screen "Dos" 800x480, template "Main"
   Group "Group_1" at 127,146 size 416x126; Text 'Мешалка 1'; PictureList "Motor"; TextList "Hand"; Picture "z2use_3"
   Group "Group_2" at 127,285 size 416x126; Text 'Мешалка 1'; PictureList "Motor"; TextList "Hand"; Picture "z2use_3"
   Rectangle "Rectangle_1" at 127,7 size 416x126
      Appearance <- "Motors_DB_M1_CMD_Sim"
   GraphicIOField "Graphic I/O field_2" at 134,43 size 43x85; PictureList "Motor"
      ProcessValue <- "Motors_DB_M1_Status"
   Button "Button_7" at 213,41 size 90x22; TextOff 'Авто'; TextList "Hand"
      on Click: InvertBit("Motors_DB_M1_CMD_Hand")
      Appearance <- "Motors_DB_M1_CMD_Hand"
      ProcessValue <- "Motors_DB_M1_CMD_Hand"
   Button "Button_8" at 258,63 size 45x22; TextOff 'Выкл'
      on Click: ResetBit("Motors_DB_M1_CMD_Start_M")
   Button "Button_9" at 213,86 size 90x20; TextOff 'Сервис'
      on Click: InvertBit("Motors_DB_M1_CMD_Service")
      Appearance <- "Motors_DB_M1_CMD_Service"
   Button "Button_13" at 213,63 size 45x22; TextOff 'Вкл'
      on Click: SetBit("Motors_DB_M1_CMD_Start_M")
      Appearance <- "Motors_DB_M1_CMD_Start_M"
   TextField "Text field_13" at 133,12 size 171x26; Text 'Дозатор 1'
   TextField "Text field_15" at 310,12 size 99x18; Text 'Ожидание ОС, с'
   GraphicView "Graphic view_1" at 180,42 size 25x25; Picture "z2use_3"
      Visibility <- "Motors_DB_M1_CMD_Hand"
   GraphicView "Graphic view_8" at 180,74 size 25x25; Picture "force"
      Visibility <- "Motors_DB_M1_CMD_Force"
   GraphicView "Graphic view_11" at 180,103 size 25x25; Picture "service"
      Visibility <- "Motors_DB_M1_CMD_Service"
   TextField "Text field_3" at 436,31 size 20x18; Text 'QF'
   TextField "Text field_10" at 436,56 size 21x18; Text 'KM'
   TextField "Text field_12" at 436,82 size 44x18; Text 'Service'
   TextField "Text field_14" at 436,108 size 41x18; Text 'Termo'
   TextField "Text field_4" at 416,10 size 120x22; Text 'Использовать:'
   Button "Button_21" at 478,32 size 60x20; TextOff 'Text'; Authorization "Operator"; PictureList "ON_OFF"
      on Click: InvertBit("Motors_DB_M1_Use_QF")
      ProcessValue <- "Motors_DB_M1_Use_QF"
   Button "Button_22" at 478,56 size 60x20; TextOff 'Text'; PictureList "ON_OFF"; Authorization "Operator"
      on Click: InvertBit("Motors_DB_M1_Use_KM")
      ProcessValue <- "Motors_DB_M1_Use_KM"
   Button "Button_24" at 478,80 size 60x20; TextOff 'Text'; PictureList "ON_OFF"; Authorization "Operator"
      on Click: InvertBit("Motors_DB_M1_Use_Serivce")
      ProcessValue <- "Motors_DB_M1_Use_Serivce"
   Button "Button_25" at 478,105 size 60x20; TextOff 'Text'; PictureList "ON_OFF"; Authorization "Operator"
      on Click: InvertBit("Motors_DB_M1_Use_Termo")
      ProcessValue <- "Motors_DB_M1_Use_Termo"
   Button "Button_26" at 416,31 size 20x20; TextOff 'Text'; Authorization "Operator"; PictureList "ok"
      ProcessValue <- "Motors_DB_M1_FB_QF"
   Button "Button_27" at 416,55 size 20x20; TextOff 'Text'; PictureList "ok"; Authorization "Operator"
      ProcessValue <- "Motors_DB_M1_FB_KM"
   Button "Button_29" at 416,80 size 20x20; TextOff 'Text'; PictureList "ok"; Authorization "Operator"
      ProcessValue <- "Motors_DB_M1_Use_Serivce"
   Button "Button_30" at 416,105 size 20x20; TextOff 'Text'; PictureList "ok"; Authorization "Operator"
      ProcessValue <- "Motors_DB_M1_FB_Termo"
   TextField "Text field_1" at 323,87 size 79x18; Text 'Наработка, ч'
   TextField "Text field_2" at 309,34 size 37x18; Text 'Старт'
   IOField "I/O field_5" at 348,32 size 30x20; FormatPattern 99
      ProcessValue <- "Motors_DB_M1_Wait_On_SP"
   IOField "I/O field_12" at 348,55 size 30x20; FormatPattern 99
      ProcessValue <- "Motors_DB_M1_Wait_Off_SP"
   TextField "Text field_5" at 309,55 size 32x18; Text 'Стоп'
   IOField "I/O field_13" at 378,32 size 30x20; FormatPattern 99
      ProcessValue <- "Motors_DB_M1_Wait_On_Now"
   IOField "I/O field_14" at 378,55 size 30x20; FormatPattern 99
      ProcessValue <- "Motors_DB_M1_Wait_Off_Now"
   IOField "I/O field_16" at 313,105 size 98x20; FormatPattern 9999999999
      ProcessValue <- "Motors_DB_M1_Res_h"
   Button "Button_11" at 213,106 size 90x20; TextOff 'Force'
      on Click: InvertBit("Motors_DB_M1_CMD_Force")
      Appearance <- "Motors_DB_M1_CMD_Force"
   Rectangle "Rectangle_4" at 550,7 size 177x126
      Appearance <- "Motors_DB_M1_CMD_Sim"
   TextField "Text field_31" at 605,8 size 68x22; Text 'Уставка'
   Button "Button_46" at 594,40 size 90x22; TextOff 'Авто'; TextList "Hand"
      on Click: InvertBit("AOx_DB_M1_SP_CMD_Hand")
      ProcessValue <- "AOx_DB_M1_SP_CMD_Hand"
      Appearance <- "AOx_DB_M1_SP_CMD_Hand"
   IOField "I/O field_15" at 594,72 size 90x20; FormatPattern 99999.99
      ProcessValue <- "AOx_DB_M1_SP_SP"
   IOField "I/O field_17" at 594,103 size 90x20; FormatPattern 99999.99
      ProcessValue <- "AOx_DB_M1_SP_SP_M"
   Rectangle "Rectangle_5" at 550,146 size 177x126
      Appearance <- "Motors_DB_M2_CMD_Sim"
   TextField "Text field_32" at 605,147 size 68x22; Text 'Уставка'
   Button "Button_47" at 594,179 size 90x22; TextOff 'Авто'; TextList "Hand"
      on Click: InvertBit("AOx_DB_M2_SP_CMD_Hand")
      Appearance <- "AOx_DB_M2_SP_CMD_Hand"
      ProcessValue <- "AOx_DB_M2_SP_CMD_Hand"
   IOField "I/O field_18" at 594,211 size 90x20; FormatPattern 99999.99
      ProcessValue <- "AOx_DB_M2_SP_SP"
   IOField "I/O field_19" at 594,242 size 90x20; FormatPattern 99999.99
      ProcessValue <- "AOx_DB_M2_SP_SP_M"
   Rectangle "Rectangle_6" at 550,285 size 177x126
      Appearance <- "Motors_DB_M3_CMD_Sim"
   TextField "Text field_33" at 605,286 size 68x22; Text 'Уставка'
   Button "Button_48" at 594,318 size 90x22; TextOff 'Авто'; TextList "Hand"
      on Click: InvertBit("AOx_DB_M3_SP_CMD_Hand")
      Appearance <- "AOx_DB_M3_SP_CMD_Hand"
      ProcessValue <- "AOx_DB_M3_SP_CMD_Hand"
   IOField "I/O field_20" at 594,350 size 90x20; FormatPattern 99999.99
      ProcessValue <- "AOx_DB_M3_SP_SP"
   IOField "I/O field_21" at 594,381 size 90x20; FormatPattern 99999.99
      ProcessValue <- "AOx_DB_M3_SP_SP_M"
   Button "Button_1" at 7,5 size 96x32; TextOff 'Насосы'; Authorization "Admin"
      on Release: ActivateScreen("Dos", 0); SetTag("settings", 1)
      Appearance <- "settings"
   Button "Button_2" at 7,51 size 96x32; TextOff 'Расход-1'; Authorization "Admin"
      on Release: ActivateScreen("Flow", 0); SetTag("settings", 2)
      Appearance <- "settings"
   Button "Button_3" at 7,140 size 96x32; TextOff 'Мутность'; Authorization "Admin"
      on Release: ActivateScreen("Trans", 0); SetTag("settings", 4)
      Appearance <- "settings"
   Button "Button_5" at 7,184 size 96x32; TextOff 'DI'; Authorization "Admin"
      on Release: ActivateScreen("DI", 0); SetTag("settings", 5)
      Appearance <- "settings"
   Button "Button_6" at 7,229 size 96x32; TextOff 'DO'; Authorization "Admin"
      on Release: ActivateScreen("DO", 0); SetTag("settings", 6)
      Appearance <- "settings"
   Button "Button_4" at 7,274 size 96x32; TextOff 'PID'; Authorization "Admin"
      on Release: ActivateScreen("PID_settings", 0); SetTag("settings", 7)
      Appearance <- "settings"
   Button "Button_49" at 7,95 size 96x32; TextOff 'Расход-2'; Authorization "Admin"
      on Release: ActivateScreen("Flow_1", 0); SetTag("settings", 3)
      Appearance <- "settings"
   Rectangle "Rectangle_2" at 127,146 size 416x126
      Appearance <- "Motors_DB_M2_CMD_Sim"
   GraphicIOField "Graphic I/O field_1" at 134,182 size 43x85; PictureList "Motor"
      ProcessValue <- "Motors_DB_M2_Status"
   Button "Button_10" at 213,180 size 90x22; TextOff 'Авто'; TextList "Hand"
      on Click: InvertBit("Motors_DB_M2_CMD_Hand")
      Appearance <- "Motors_DB_M2_CMD_Hand"
      ProcessValue <- "Motors_DB_M2_CMD_Hand"
   Button "Button_12" at 258,202 size 45x22; TextOff 'Выкл'
      on Click: ResetBit("Motors_DB_M2_CMD_Start_M")
   Button "Button_14" at 213,225 size 90x20; TextOff 'Сервис'
      on Click: InvertBit("Motors_DB_M2_CMD_Service")
      Appearance <- "Motors_DB_M2_CMD_Service"
   Button "Button_15" at 213,202 size 45x22; TextOff 'Вкл'
      on Click: SetBit("Motors_DB_M2_CMD_Start_M")
      Appearance <- "Motors_DB_M2_CMD_Start_M"
   TextField "Text field_6" at 133,151 size 171x26; Text 'Дозатор 2'
   TextField "Text field_7" at 310,151 size 99x18; Text 'Ожидание ОС, с'
   GraphicView "Graphic view_2" at 180,181 size 25x25; Picture "z2use_3"
      Visibility <- "Motors_DB_M2_CMD_Hand"
   GraphicView "Graphic view_3" at 180,213 size 25x25; Picture "force"
      Visibility <- "Motors_DB_M2_CMD_Force"
   GraphicView "Graphic view_4" at 180,242 size 25x25; Picture "service"
      Visibility <- "Motors_DB_M2_CMD_Service"
   TextField "Text field_8" at 436,170 size 20x18; Text 'QF'
   TextField "Text field_9" at 436,195 size 21x18; Text 'KM'
   TextField "Text field_11" at 436,221 size 44x18; Text 'Service'
   TextField "Text field_16" at 436,247 size 41x18; Text 'Termo'
   TextField "Text field_17" at 416,149 size 120x22; Text 'Использовать:'
   Button "Button_16" at 478,171 size 60x20; TextOff 'Text'; PictureList "ON_OFF"; Authorization "Operator"
      on Click: InvertBit("Motors_DB_M2_Use_QF")
      ProcessValue <- "Motors_DB_M2_Use_QF"
   Button "Button_17" at 478,195 size 60x20; TextOff 'Text'; Authorization "Operator"; PictureList "ON_OFF"
      on Click: InvertBit("Motors_DB_M2_Use_KM")
      ProcessValue <- "Motors_DB_M2_Use_KM"
   Button "Button_18" at 478,219 size 60x20; TextOff 'Text'; Authorization "Operator"; PictureList "ON_OFF"
      on Click: InvertBit("Motors_DB_M2_Use_Serivce")
      ProcessValue <- "Motors_DB_M2_Use_Serivce"
   Button "Button_19" at 478,244 size 60x20; TextOff 'Text'; Authorization "Operator"; PictureList "ON_OFF"
      on Click: InvertBit("Motors_DB_M2_Use_Termo")
      ProcessValue <- "Motors_DB_M2_Use_Termo"
   Button "Button_20" at 416,170 size 20x20; TextOff 'Text'; PictureList "ok"; Authorization "Operator"
      ProcessValue <- "Motors_DB_M2_FB_QF"
   Button "Button_23" at 416,194 size 20x20; TextOff 'Text'; Authorization "Operator"; PictureList "ok"
      ProcessValue <- "Motors_DB_M2_FB_KM"
   Button "Button_28" at 416,219 size 20x20; TextOff 'Text'; Authorization "Operator"; PictureList "ok"
      ProcessValue <- "Motors_DB_M2_Use_Serivce"
   Button "Button_31" at 416,244 size 20x20; TextOff 'Text'; Authorization "Operator"; PictureList "ok"
      ProcessValue <- "Motors_DB_M2_FB_Termo"
   TextField "Text field_18" at 323,226 size 79x18; Text 'Наработка, ч'
   TextField "Text field_19" at 309,173 size 37x18; Text 'Старт'
   IOField "I/O field_1" at 348,171 size 30x20; FormatPattern 99
      ProcessValue <- "Motors_DB_M2_Wait_On_SP"
   IOField "I/O field_2" at 348,194 size 30x20; FormatPattern 99
      ProcessValue <- "Motors_DB_M2_Wait_Off_SP"
   TextField "Text field_20" at 309,194 size 32x18; Text 'Стоп'
   IOField "I/O field_3" at 378,171 size 30x20; FormatPattern 99
      ProcessValue <- "Motors_DB_M2_Wait_On_Now"
   IOField "I/O field_4" at 378,194 size 30x20; FormatPattern 99
      ProcessValue <- "Motors_DB_M2_Wait_Off_Now"
   IOField "I/O field_6" at 313,244 size 98x20; FormatPattern 9999999999
      ProcessValue <- "Motors_DB_M2_Res_h"
   Button "Button_32" at 213,245 size 90x20; TextOff 'Force'
      on Click: InvertBit("Motors_DB_M2_CMD_Force")
      Appearance <- "Motors_DB_M2_CMD_Force"
   Rectangle "Rectangle_3" at 127,285 size 416x126
      Appearance <- "Motors_DB_M3_CMD_Sim"
   GraphicIOField "Graphic I/O field_3" at 134,321 size 43x85; PictureList "Motor"
      ProcessValue <- "Motors_DB_M3_Status"
   Button "Button_33" at 213,319 size 90x22; TextOff 'Авто'; TextList "Hand"
      on Click: InvertBit("Motors_DB_M3_CMD_Hand")
      Appearance <- "Motors_DB_M3_CMD_Hand"
      ProcessValue <- "Motors_DB_M3_CMD_Hand"
   Button "Button_34" at 258,341 size 45x22; TextOff 'Выкл'
      on Click: ResetBit("Motors_DB_M3_CMD_Start_M")
   Button "Button_35" at 213,364 size 90x20; TextOff 'Сервис'
      on Click: InvertBit("Motors_DB_M3_CMD_Service")
      Appearance <- "Motors_DB_M3_CMD_Service"
   Button "Button_36" at 213,341 size 45x22; TextOff 'Вкл'
      on Click: SetBit("Motors_DB_M3_CMD_Start_M")
      Appearance <- "Motors_DB_M3_CMD_Start_M"
   TextField "Text field_21" at 133,290 size 171x26; Text 'Дозатор 3'
   TextField "Text field_22" at 310,290 size 99x18; Text 'Ожидание ОС, с'
   GraphicView "Graphic view_5" at 180,320 size 25x25; Picture "z2use_3"
      Visibility <- "Motors_DB_M3_CMD_Hand"
   GraphicView "Graphic view_6" at 180,352 size 25x25; Picture "force"
      Visibility <- "Motors_DB_M3_CMD_Force"
   GraphicView "Graphic view_7" at 180,381 size 25x25; Picture "service"
      Visibility <- "Motors_DB_M3_CMD_Service"
   TextField "Text field_23" at 436,309 size 20x18; Text 'QF'
   TextField "Text field_24" at 436,334 size 21x18; Text 'KM'
   TextField "Text field_25" at 436,360 size 44x18; Text 'Service'
   TextField "Text field_26" at 436,386 size 41x18; Text 'Termo'
   TextField "Text field_27" at 416,288 size 120x22; Text 'Использовать:'
   Button "Button_37" at 478,310 size 60x20; TextOff 'Text'; PictureList "ON_OFF"; Authorization "Operator"
      on Click: InvertBit("Motors_DB_M3_Use_QF")
      ProcessValue <- "Motors_DB_M3_Use_QF"
   Button "Button_38" at 478,334 size 60x20; TextOff 'Text'; Authorization "Operator"; PictureList "ON_OFF"
      on Click: InvertBit("Motors_DB_M3_Use_KM")
      ProcessValue <- "Motors_DB_M3_Use_KM"
   Button "Button_39" at 478,358 size 60x20; TextOff 'Text'; Authorization "Operator"; PictureList "ON_OFF"
      on Click: InvertBit("Motors_DB_M3_Use_Serivce")
      ProcessValue <- "Motors_DB_M3_Use_Serivce"
   Button "Button_40" at 478,383 size 60x20; TextOff 'Text'; Authorization "Operator"; PictureList "ON_OFF"
      on Click: InvertBit("Motors_DB_M3_Use_Termo")
      ProcessValue <- "Motors_DB_M3_Use_Termo"
   Button "Button_41" at 416,309 size 20x20; TextOff 'Text'; PictureList "ok"; Authorization "Operator"
      ProcessValue <- "Motors_DB_M3_FB_QF"
   Button "Button_42" at 416,333 size 20x20; TextOff 'Text'; Authorization "Operator"; PictureList "ok"
      ProcessValue <- "Motors_DB_M3_FB_KM"
   Button "Button_43" at 416,358 size 20x20; TextOff 'Text'; Authorization "Operator"; PictureList "ok"
      ProcessValue <- "Motors_DB_M3_Use_Serivce"
   Button "Button_44" at 416,383 size 20x20; TextOff 'Text'; Authorization "Operator"; PictureList "ok"
      ProcessValue <- "Motors_DB_M3_FB_Termo"
   TextField "Text field_28" at 323,365 size 79x18; Text 'Наработка, ч'
   TextField "Text field_29" at 309,312 size 37x18; Text 'Старт'
   IOField "I/O field_7" at 348,310 size 30x20; FormatPattern 99
      ProcessValue <- "Motors_DB_M3_Wait_On_SP"
   IOField "I/O field_8" at 348,333 size 30x20; FormatPattern 99
      ProcessValue <- "Motors_DB_M3_Wait_Off_SP"
   TextField "Text field_30" at 309,333 size 32x18; Text 'Стоп'
   IOField "I/O field_9" at 378,310 size 30x20; FormatPattern 99
      ProcessValue <- "Motors_DB_M3_Wait_On_Now"
   IOField "I/O field_10" at 378,333 size 30x20; FormatPattern 99
      ProcessValue <- "Motors_DB_M3_Wait_Off_Now"
   IOField "I/O field_11" at 313,383 size 98x20; FormatPattern 9999999999
      ProcessValue <- "Motors_DB_M3_Res_h"
   Button "Button_45" at 213,384 size 90x20; TextOff 'Force'
      on Click: InvertBit("Motors_DB_M3_CMD_Force")
      Appearance <- "Motors_DB_M3_CMD_Force"

screen "Trans" 800x480, template "Main"
   TextField "Text field_2" at 210,15 size 67x22; Text 'Датчик:'
   TextField "Text field_4" at 273,15 size 94x22; Text 'Мутность 1'
   TextField "Text field_7" at 390,18 size 43x22; Text 'вход'
   TextField "Text field_8" at 390,43 size 56x22; Text 'выход'
   IOField "I/O field_1" at 452,19 size 102x26; FormatPattern s99999.99
      ProcessValue <- "AIx_DB_Trans_1_Converter_Min_In"
   IOField "I/O field_2" at 452,41 size 102x26; FormatPattern s99999.99
      ProcessValue <- "AIx_DB_Trans_1_Converter_Min_Out"
   IOField "I/O field_3" at 551,19 size 102x26; FormatPattern s99999.99
      ProcessValue <- "AIx_DB_Trans_1_Converter_Max_In"
   IOField "I/O field_4" at 551,41 size 102x26; FormatPattern s99999.99
      ProcessValue <- "AIx_DB_Trans_1_Converter_Max_Out"
   TextField "Text field_9" at 389,68 size 101x22; Text 'Фильтрация'
   TextField "Text field_10" at 390,96 size 36x22; Text 'RTD'
   Button "Button_7" at 489,71 size 20x20; TextOff 'Text'; PictureList "ok"
      on Click: InvertBit("AIx_DB_Trans_1_Use_Filter")
      ProcessValue <- "AIx_DB_Trans_1_Use_Filter"
   Button "Button_8" at 489,96 size 20x20; TextOff 'Text'; PictureList "ok"
      on Click: InvertBit("AIx_DB_Trans_1_Use_RTD")
      ProcessValue <- "AIx_DB_Trans_1_Use_RTD"
   IOField "I/O field_5" at 516,68 size 65x25; FormatPattern 999
      ProcessValue <- "AIx_DB_Trans_1_Filter_SP"
   IOField "I/O field_6" at 516,93 size 65x25; FormatPattern 999
      ProcessValue <- "AIx_DB_Trans_1_RTD_c"
   TextField "Text field_11" at 210,36 size 79x22; Text 'Поправка'
   IOField "I/O field_7" at 293,36 size 78x23; FormatPattern s999.9
      ProcessValue <- "AIx_DB_Trans_1_Calibration"
   Button "Button_9" at 396,176 size 248x28; TextOff 'Use'
      on Click: InvertBit("AIx_DB_Trans_1_CMD_Start_A")
      Appearance <- "AIx_DB_Trans_1_CMD_Start_A"
   Button "Button_10" at 213,66 size 68x28; TextOff 'Hand'
      on Click: InvertBit("AIx_DB_Trans_1_CMD_Hand")
      Appearance <- "AIx_DB_Trans_1_CMD_Hand"
   IOField "I/O field_8" at 293,66 size 78x28; FormatPattern s9999.9
      ProcessValue <- "AIx_DB_Trans_1_Result"
   TextField "Text field_12" at 436,123 size 27x22; Text 'NC'
   TextField "Text field_13" at 437,143 size 25x22; Text 'SC'
   TextField "Text field_14" at 210,125 size 27x22; Text 'HH'
   TextField "Text field_15" at 216,145 size 16x22; Text 'H'
   TextField "Text field_16" at 217,165 size 14x22; Text 'L'
   TextField "Text field_17" at 212,186 size 23x22; Text 'LL'
   IOField "I/O field_11" at 472,123 size 58x21; FormatPattern s99999
      ProcessValue <- "AIx_DB_Trans_1_SP_NC"
   IOField "I/O field_12" at 472,143 size 58x21; FormatPattern s99999
      ProcessValue <- "AIx_DB_Trans_1_SP_SC"
   IOField "I/O field_13" at 246,125 size 58x21; FormatPattern 99999
      ProcessValue <- "AIx_DB_Trans_1_SP_HH"
   IOField "I/O field_14" at 246,145 size 58x21; FormatPattern 99999
      ProcessValue <- "AIx_DB_Trans_1_SP_H"
   IOField "I/O field_15" at 246,165 size 58x21; FormatPattern s99999
      ProcessValue <- "AIx_DB_Trans_1_SP_L"
   IOField "I/O field_16" at 246,185 size 58x21; FormatPattern s99999
      ProcessValue <- "AIx_DB_Trans_1_SP_LL"
   IOField "I/O field_17" at 546,123 size 58x21; FormatPattern 999
      ProcessValue <- "AIx_DB_Trans_1_Timers_NC_SP"
   IOField "I/O field_18" at 546,143 size 58x21; FormatPattern 999
      ProcessValue <- "AIx_DB_Trans_1_Timers_SC_SP"
   IOField "I/O field_19" at 320,125 size 58x21; FormatPattern 999
      ProcessValue <- "AIx_DB_Trans_1_Timers_HH_SP"
   IOField "I/O field_20" at 320,145 size 58x21; FormatPattern 999
      ProcessValue <- "AIx_DB_Trans_1_Timers_H_SP"
   IOField "I/O field_21" at 320,165 size 58x21; FormatPattern 999
      ProcessValue <- "AIx_DB_Trans_1_Timers_L_SP"
   IOField "I/O field_22" at 320,185 size 58x21; FormatPattern 999
      ProcessValue <- "AIx_DB_Trans_1_Timers_LL_SP"
   IOField "I/O field_23" at 582,93 size 65x25; FormatPattern s99999
      ProcessValue <- "AIx_DB_Trans_1_Signal"
   TextField "Text field_18" at 210,97 size 68x22; Text 'Уставка'
   TextField "Text field_19" at 299,97 size 79x22; Text 'Время (с)'
   TextField "Text field_1" at 214,248 size 67x22; Text 'Датчик:'
   TextField "Text field_3" at 277,248 size 94x22; Text 'Мутность 2'
   TextField "Text field_5" at 394,251 size 43x22; Text 'вход'
   TextField "Text field_6" at 394,276 size 56x22; Text 'выход'
   IOField "I/O field_9" at 456,252 size 102x26; FormatPattern s99999.99
      ProcessValue <- "AIx_DB_Trans_2_Converter_Min_In"
   IOField "I/O field_10" at 456,274 size 102x26; FormatPattern s99999.99
      ProcessValue <- "AIx_DB_Trans_2_Converter_Min_Out"
   IOField "I/O field_24" at 555,252 size 102x26; FormatPattern s99999.99
      ProcessValue <- "AIx_DB_Trans_2_Converter_Max_In"
   IOField "I/O field_25" at 555,274 size 102x26; FormatPattern s99999.99
      ProcessValue <- "AIx_DB_Trans_2_Converter_Max_Out"
   TextField "Text field_20" at 393,301 size 101x22; Text 'Фильтрация'
   TextField "Text field_21" at 394,329 size 36x22; Text 'RTD'
   Button "Button_11" at 493,304 size 20x20; TextOff 'Text'; PictureList "ok"
      on Click: InvertBit("AIx_DB_Trans_2_Use_Filter")
      ProcessValue <- "AIx_DB_Trans_2_Use_Filter"
   Button "Button_12" at 493,329 size 20x20; TextOff 'Text'; PictureList "ok"
      on Click: InvertBit("AIx_DB_Trans_2_Use_RTD")
      ProcessValue <- "AIx_DB_Trans_2_Use_RTD"
   IOField "I/O field_26" at 520,301 size 65x25; FormatPattern 999
      ProcessValue <- "AIx_DB_Trans_2_Filter_SP"
   IOField "I/O field_27" at 520,326 size 65x25; FormatPattern 999
      ProcessValue <- "AIx_DB_Trans_2_RTD_c"
   TextField "Text field_22" at 214,269 size 79x22; Text 'Поправка'
   IOField "I/O field_28" at 297,269 size 78x23; FormatPattern s999.9
      ProcessValue <- "AIx_DB_Trans_2_Calibration"
   Button "Button_13" at 400,409 size 248x28; TextOff 'Use'
      on Click: InvertBit("AIx_DB_Trans_2_CMD_Start_A")
      Appearance <- "AIx_DB_Trans_2_CMD_Start_A"
   Button "Button_14" at 217,299 size 68x28; TextOff 'Hand'
      on Click: InvertBit("AIx_DB_Trans_2_CMD_Hand")
      Appearance <- "AIx_DB_Trans_2_CMD_Hand"
   IOField "I/O field_29" at 297,299 size 78x28; FormatPattern s9999.9
      ProcessValue <- "AIx_DB_Trans_2_Result"
   TextField "Text field_23" at 440,356 size 27x22; Text 'NC'
   TextField "Text field_24" at 441,376 size 25x22; Text 'SC'
   TextField "Text field_25" at 214,358 size 27x22; Text 'HH'
   TextField "Text field_26" at 220,378 size 16x22; Text 'H'
   TextField "Text field_27" at 221,398 size 14x22; Text 'L'
   TextField "Text field_28" at 216,419 size 23x22; Text 'LL'
   IOField "I/O field_30" at 476,356 size 58x21; FormatPattern s99999
      ProcessValue <- "AIx_DB_Trans_2_SP_NC"
   IOField "I/O field_31" at 476,376 size 58x21; FormatPattern s99999
      ProcessValue <- "AIx_DB_Trans_2_SP_SC"
   IOField "I/O field_32" at 250,358 size 58x21; FormatPattern 99999
      ProcessValue <- "AIx_DB_Trans_2_SP_HH"
   IOField "I/O field_33" at 250,378 size 58x21; FormatPattern 99999
      ProcessValue <- "AIx_DB_Trans_2_SP_H"
   IOField "I/O field_34" at 250,398 size 58x21; FormatPattern s99999
      ProcessValue <- "AIx_DB_Trans_2_SP_L"
   IOField "I/O field_35" at 250,418 size 58x21; FormatPattern s99999
      ProcessValue <- "AIx_DB_Trans_2_SP_LL"
   IOField "I/O field_36" at 550,356 size 58x21; FormatPattern 999
      ProcessValue <- "AIx_DB_Trans_2_Timers_NC_SP"
   IOField "I/O field_37" at 550,376 size 58x21; FormatPattern 999
      ProcessValue <- "AIx_DB_Trans_2_Timers_SC_SP"
   IOField "I/O field_38" at 324,358 size 58x21; FormatPattern 999
      ProcessValue <- "AIx_DB_Trans_2_Timers_HH_SP"
   IOField "I/O field_39" at 324,378 size 58x21; FormatPattern 999
      ProcessValue <- "AIx_DB_Trans_2_Timers_H_SP"
   IOField "I/O field_40" at 324,398 size 58x21; FormatPattern 999
      ProcessValue <- "AIx_DB_Trans_2_Timers_L_SP"
   IOField "I/O field_41" at 324,418 size 58x21; FormatPattern 999
      ProcessValue <- "AIx_DB_Trans_2_Timers_LL_SP"
   IOField "I/O field_42" at 586,326 size 65x25; FormatPattern s99999
      ProcessValue <- "AIx_DB_Trans_2_Signal"
   TextField "Text field_29" at 214,330 size 68x22; Text 'Уставка'
   TextField "Text field_30" at 303,330 size 79x22; Text 'Время (с)'
   Button "Button_1" at 7,5 size 96x32; TextOff 'Насосы'; Authorization "Admin"
      on Release: ActivateScreen("Dos", 0); SetTag("settings", 1)
      Appearance <- "settings"
   Button "Button_2" at 7,51 size 96x32; TextOff 'Расход-1'; Authorization "Admin"
      on Release: ActivateScreen("Flow", 0); SetTag("settings", 2)
      Appearance <- "settings"
   Button "Button_3" at 7,140 size 96x32; TextOff 'Мутность'; Authorization "Admin"
      on Release: ActivateScreen("Trans", 0); SetTag("settings", 4)
      Appearance <- "settings"
   Button "Button_5" at 7,184 size 96x32; TextOff 'DI'; Authorization "Admin"
      on Release: ActivateScreen("DI", 0); SetTag("settings", 5)
      Appearance <- "settings"
   Button "Button_6" at 7,229 size 96x32; TextOff 'DO'; Authorization "Admin"
      on Release: ActivateScreen("DO", 0); SetTag("settings", 6)
      Appearance <- "settings"
   Button "Button_4" at 7,274 size 96x32; TextOff 'PID'; Authorization "Admin"
      on Release: ActivateScreen("PID_settings", 0); SetTag("settings", 7)
      Appearance <- "settings"
   Button "Button_15" at 7,95 size 96x32; TextOff 'Расход-2'; Authorization "Admin"
      on Release: ActivateScreen("Flow_1", 0); SetTag("settings", 3)
      Appearance <- "settings"

screen "Flow" 800x480, template "Main"
   TextField "Text field_2" at 210,15 size 67x22; Text 'Датчик:'
   TextField "Text field_4" at 273,15 size 113x22; Text 'Расходомер 1'
   TextField "Text field_7" at 390,18 size 43x22; Text 'вход'
   TextField "Text field_8" at 390,43 size 56x22; Text 'выход'
   IOField "I/O field_1" at 452,19 size 102x26; FormatPattern s99999.99
      ProcessValue <- "AIx_DB_Flow_1_Converter_Min_In"
   IOField "I/O field_2" at 452,41 size 102x26; FormatPattern s99999.99
      ProcessValue <- "AIx_DB_Flow_1_Converter_Min_Out"
   IOField "I/O field_3" at 551,19 size 102x26; FormatPattern s99999.99
      ProcessValue <- "AIx_DB_Flow_1_Converter_Max_In"
   IOField "I/O field_4" at 551,41 size 102x26; FormatPattern s99999.99
      ProcessValue <- "AIx_DB_Flow_1_Converter_Max_Out"
   TextField "Text field_9" at 389,68 size 101x22; Text 'Фильтрация'
   TextField "Text field_10" at 390,96 size 36x22; Text 'RTD'
   Button "Button_7" at 489,71 size 20x20; TextOff 'Text'; PictureList "ok"
      on Click: InvertBit("AIx_DB_Flow_1_Use_Filter")
      ProcessValue <- "AIx_DB_Flow_1_Use_Filter"
   Button "Button_8" at 489,96 size 20x20; TextOff 'Text'; PictureList "ok"
      on Click: InvertBit("AIx_DB_Flow_1_Use_RTD")
      ProcessValue <- "AIx_DB_Flow_1_Use_RTD"
   IOField "I/O field_5" at 516,68 size 65x25; FormatPattern 999
      ProcessValue <- "AIx_DB_Flow_1_Filter_SP"
   IOField "I/O field_6" at 516,93 size 65x25; FormatPattern 999
      ProcessValue <- "AIx_DB_Flow_1_RTD_c"
   TextField "Text field_11" at 210,36 size 79x22; Text 'Поправка'
   IOField "I/O field_7" at 293,36 size 78x23; FormatPattern s999.9
      ProcessValue <- "AIx_DB_Flow_1_Calibration"
   Button "Button_9" at 396,176 size 248x28; TextOff 'Use'
      on Click: InvertBit("AIx_DB_Flow_1_CMD_Start_A")
      Appearance <- "AIx_DB_Flow_1_CMD_Start_A"
   Button "Button_10" at 213,66 size 68x28; TextOff 'Hand'
      on Click: InvertBit("AIx_DB_Flow_1_CMD_Hand")
      Appearance <- "AIx_DB_Flow_1_CMD_Hand"
   IOField "I/O field_8" at 293,66 size 78x28; FormatPattern s9999.9
      ProcessValue <- "AIx_DB_Flow_1_Result"
   TextField "Text field_12" at 436,123 size 27x22; Text 'NC'
   TextField "Text field_13" at 437,143 size 25x22; Text 'SC'
   TextField "Text field_14" at 210,125 size 27x22; Text 'HH'
   TextField "Text field_15" at 216,145 size 16x22; Text 'H'
   TextField "Text field_16" at 217,165 size 14x22; Text 'L'
   TextField "Text field_17" at 212,186 size 23x22; Text 'LL'
   IOField "I/O field_11" at 472,123 size 58x21; FormatPattern s99999
      ProcessValue <- "AIx_DB_Flow_1_SP_NC"
   IOField "I/O field_12" at 472,143 size 58x21; FormatPattern s99999
      ProcessValue <- "AIx_DB_Flow_1_SP_SC"
   IOField "I/O field_13" at 246,125 size 58x21; FormatPattern 99999
      ProcessValue <- "AIx_DB_Flow_1_SP_HH"
   IOField "I/O field_14" at 246,145 size 58x21; FormatPattern 99999
      ProcessValue <- "AIx_DB_Flow_1_SP_H"
   IOField "I/O field_15" at 246,165 size 58x21; FormatPattern s99999
      ProcessValue <- "AIx_DB_Flow_1_SP_L"
   IOField "I/O field_16" at 246,185 size 58x21; FormatPattern s99999
      ProcessValue <- "AIx_DB_Flow_1_SP_LL"
   IOField "I/O field_17" at 546,123 size 58x21; FormatPattern 999
      ProcessValue <- "AIx_DB_Flow_1_Timers_NC_SP"
   IOField "I/O field_18" at 546,143 size 58x21; FormatPattern 999
      ProcessValue <- "AIx_DB_Flow_1_Timers_SC_SP"
   IOField "I/O field_19" at 320,125 size 58x21; FormatPattern 999
      ProcessValue <- "AIx_DB_Flow_1_Timers_HH_SP"
   IOField "I/O field_20" at 320,145 size 58x21; FormatPattern 999
      ProcessValue <- "AIx_DB_Flow_1_Timers_H_SP"
   IOField "I/O field_21" at 320,165 size 58x21; FormatPattern 999
      ProcessValue <- "AIx_DB_Flow_1_Timers_L_SP"
   IOField "I/O field_22" at 320,185 size 58x21; FormatPattern 999
      ProcessValue <- "AIx_DB_Flow_1_Timers_LL_SP"
   IOField "I/O field_23" at 582,93 size 65x25; FormatPattern s99999
      ProcessValue <- "AIx_DB_Flow_1_Signal"
   TextField "Text field_18" at 210,97 size 68x22; Text 'Уставка'
   TextField "Text field_19" at 299,97 size 79x22; Text 'Время (с)'
   TextField "Text field_1" at 214,248 size 67x22; Text 'Датчик:'
   TextField "Text field_3" at 277,248 size 113x22; Text 'Расходомер 2'
   TextField "Text field_5" at 394,251 size 43x22; Text 'вход'
   TextField "Text field_6" at 394,276 size 56x22; Text 'выход'
   IOField "I/O field_9" at 456,252 size 102x26; FormatPattern s99999.99
      ProcessValue <- "AIx_DB_Flow_2_Converter_Min_In"
   IOField "I/O field_10" at 456,274 size 102x26; FormatPattern s99999.99
      ProcessValue <- "AIx_DB_Flow_2_Converter_Min_Out"
   IOField "I/O field_24" at 555,252 size 102x26; FormatPattern s99999.99
      ProcessValue <- "AIx_DB_Flow_2_Converter_Max_In"
   IOField "I/O field_25" at 555,274 size 102x26; FormatPattern s99999.99
      ProcessValue <- "AIx_DB_Flow_2_Converter_Max_Out"
   TextField "Text field_20" at 393,301 size 101x22; Text 'Фильтрация'
   TextField "Text field_21" at 394,329 size 36x22; Text 'RTD'
   Button "Button_11" at 493,304 size 20x20; TextOff 'Text'; PictureList "ok"
      on Click: InvertBit("AIx_DB_Flow_2_Use_Filter")
      ProcessValue <- "AIx_DB_Flow_2_Use_Filter"
   Button "Button_12" at 493,329 size 20x20; TextOff 'Text'; PictureList "ok"
      on Click: InvertBit("AIx_DB_Flow_2_Use_RTD")
      ProcessValue <- "AIx_DB_Flow_2_Use_RTD"
   IOField "I/O field_26" at 520,301 size 65x25; FormatPattern 999
      ProcessValue <- "AIx_DB_Flow_2_Filter_SP"
   IOField "I/O field_27" at 520,326 size 65x25; FormatPattern 999
      ProcessValue <- "AIx_DB_Flow_2_RTD_c"
   TextField "Text field_22" at 214,269 size 79x22; Text 'Поправка'
   IOField "I/O field_28" at 297,269 size 78x23; FormatPattern s999.9
      ProcessValue <- "AIx_DB_Flow_2_Calibration"
   Button "Button_13" at 400,409 size 248x28; TextOff 'Use'
      on Click: InvertBit("AIx_DB_Flow_2_CMD_Start_A")
      Appearance <- "AIx_DB_Flow_2_CMD_Start_A"
   Button "Button_14" at 217,299 size 68x28; TextOff 'Hand'
      on Click: InvertBit("AIx_DB_Flow_2_CMD_Hand")
      Appearance <- "AIx_DB_Flow_2_CMD_Hand"
   IOField "I/O field_29" at 297,299 size 78x28; FormatPattern s9999.9
      ProcessValue <- "AIx_DB_Flow_2_Result"
   TextField "Text field_23" at 440,356 size 27x22; Text 'NC'
   TextField "Text field_24" at 441,376 size 25x22; Text 'SC'
   TextField "Text field_25" at 214,358 size 27x22; Text 'HH'
   TextField "Text field_26" at 220,378 size 16x22; Text 'H'
   TextField "Text field_27" at 221,398 size 14x22; Text 'L'
   TextField "Text field_28" at 216,419 size 23x22; Text 'LL'
   IOField "I/O field_30" at 476,356 size 58x21; FormatPattern s99999
      ProcessValue <- "AIx_DB_Flow_2_SP_NC"
   IOField "I/O field_31" at 476,376 size 58x21; FormatPattern s99999
      ProcessValue <- "AIx_DB_Flow_2_SP_SC"
   IOField "I/O field_32" at 250,358 size 58x21; FormatPattern 99999
      ProcessValue <- "AIx_DB_Flow_2_SP_HH"
   IOField "I/O field_33" at 250,378 size 58x21; FormatPattern 99999
      ProcessValue <- "AIx_DB_Flow_2_SP_H"
   IOField "I/O field_34" at 250,398 size 58x21; FormatPattern s99999
      ProcessValue <- "AIx_DB_Flow_2_SP_L"
   IOField "I/O field_35" at 250,418 size 58x21; FormatPattern s99999
      ProcessValue <- "AIx_DB_Flow_2_SP_LL"
   IOField "I/O field_36" at 550,356 size 58x21; FormatPattern 999
      ProcessValue <- "AIx_DB_Flow_2_Timers_NC_SP"
   IOField "I/O field_37" at 550,376 size 58x21; FormatPattern 999
      ProcessValue <- "AIx_DB_Flow_2_Timers_SC_SP"
   IOField "I/O field_38" at 324,358 size 58x21; FormatPattern 999
      ProcessValue <- "AIx_DB_Flow_2_Timers_HH_SP"
   IOField "I/O field_39" at 324,378 size 58x21; FormatPattern 999
      ProcessValue <- "AIx_DB_Flow_2_Timers_H_SP"
   IOField "I/O field_40" at 324,398 size 58x21; FormatPattern 999
      ProcessValue <- "AIx_DB_Flow_2_Timers_L_SP"
   IOField "I/O field_41" at 324,418 size 58x21; FormatPattern 999
      ProcessValue <- "AIx_DB_Flow_2_Timers_LL_SP"
   IOField "I/O field_42" at 586,326 size 65x25; FormatPattern s99999
      ProcessValue <- "AIx_DB_Flow_2_Signal"
   TextField "Text field_29" at 214,330 size 68x22; Text 'Уставка'
   TextField "Text field_30" at 303,330 size 79x22; Text 'Время (с)'
   Button "Button_1" at 7,5 size 96x32; TextOff 'Насосы'; Authorization "Admin"
      on Release: ActivateScreen("Dos", 0); SetTag("settings", 1)
      Appearance <- "settings"
   Button "Button_2" at 7,51 size 96x32; TextOff 'Расход-1'; Authorization "Admin"
      on Release: ActivateScreen("Flow", 0); SetTag("settings", 2)
      Appearance <- "settings"
   Button "Button_3" at 7,140 size 96x32; TextOff 'Мутность'; Authorization "Admin"
      on Release: ActivateScreen("Trans", 0); SetTag("settings", 4)
      Appearance <- "settings"
   Button "Button_5" at 7,184 size 96x32; TextOff 'DI'; Authorization "Admin"
      on Release: ActivateScreen("DI", 0); SetTag("settings", 5)
      Appearance <- "settings"
   Button "Button_6" at 7,229 size 96x32; TextOff 'DO'; Authorization "Admin"
      on Release: ActivateScreen("DO", 0); SetTag("settings", 6)
      Appearance <- "settings"
   Button "Button_4" at 7,274 size 96x32; TextOff 'PID'; Authorization "Admin"
      on Release: ActivateScreen("PID_settings", 0); SetTag("settings", 7)
      Appearance <- "settings"
   Button "Button_15" at 7,95 size 96x32; TextOff 'Расход-2'; Authorization "Admin"
      on Release: ActivateScreen("Flow_1", 0); SetTag("settings", 3)
      Appearance <- "settings"

screen "DI" 800x480, template "Main"
   Group "Group" at 127,7 size 283x51; TextList "Hand"
   Group "Group_1" at 127,66 size 283x51; TextList "Hand"
   Group "Group_2" at 127,125 size 283x51; TextList "Hand"
   Group "Group_3" at 127,184 size 283x51; TextList "Hand"
   Group "Group_4" at 127,244 size 283x51; TextList "Hand"
   Group "Group_5" at 127,303 size 283x51; TextList "Hand"
   Group "Group_6" at 127,362 size 283x51; TextList "Hand"
   Group "Group_7" at 127,422 size 283x51; TextList "Hand"
   Group "Group_8" at 433,7 size 283x51; TextList "Hand"
   Group "Group_9" at 433,66 size 283x51; TextList "Hand"
   Button "Button_1" at 7,5 size 96x32; TextOff 'Насосы'; Authorization "Admin"
      on Release: ActivateScreen("Dos", 0); SetTag("settings", 1)
      Appearance <- "settings"
   Button "Button_2" at 7,51 size 96x32; TextOff 'Расход-1'; Authorization "Admin"
      on Release: ActivateScreen("Flow", 0); SetTag("settings", 2)
      Appearance <- "settings"
   Button "Button_3" at 7,140 size 96x32; TextOff 'Мутность'; Authorization "Admin"
      on Release: ActivateScreen("Trans", 0); SetTag("settings", 4)
      Appearance <- "settings"
   Button "Button_5" at 7,184 size 96x32; TextOff 'DI'; Authorization "Admin"
      on Release: ActivateScreen("DI", 0); SetTag("settings", 5)
      Appearance <- "settings"
   Button "Button_6" at 7,229 size 96x32; TextOff 'DO'; Authorization "Admin"
      on Release: ActivateScreen("DO", 0); SetTag("settings", 6)
      Appearance <- "settings"
   Button "Button_4" at 7,274 size 96x32; TextOff 'PID'; Authorization "Admin"
      on Release: ActivateScreen("PID_settings", 0); SetTag("settings", 7)
      Appearance <- "settings"
   Button "Button_47" at 7,95 size 96x32; TextOff 'Расход-2'; Authorization "Admin"
      on Release: ActivateScreen("Flow_1", 0); SetTag("settings", 3)
      Appearance <- "settings"
   TextField "Text field_1" at 131,10 size 45x22; Text 'I 0.0'
   TextField "Text field_2" at 176,10 size 120x22; Text 'M1 Готовность'
   Circle "Circle_1" at 131,33 size 22x22
      Appearance <- "DIx_DB_M1_QF_Input"
   Circle "Circle_2" at 154,33 size 22x22
      Appearance <- "DIx_DB_M1_QF_Signal"
   Button "Button_7" at 298,11 size 59x44; TextOff 'Авто'; TextList "Hand"
      on Click: InvertBit("DIx_DB_M1_QF_Hand")
      Appearance <- "DIx_DB_M1_QF_Hand"
      ProcessValue <- "DIx_DB_M1_QF_Hand"
   Button "Button_8" at 240,33 size 49x22; TextOff 'Выкл'
      on Click: ResetBit("DIx_DB_M1_QF_Start_M")
   Button "Button_12" at 184,33 size 47x22; TextOff 'Вкл'
      on Click: SetBit("DIx_DB_M1_QF_Start_M")
      Appearance <- "DIx_DB_M1_QF_Start_M"
   IOField "I/O field_6" at 360,33 size 23x22; FormatPattern 99
      ProcessValue <- "DIx_DB_M1_QF_Filter_On_SP"
   IOField "I/O field_7" at 383,33 size 23x22; FormatPattern 99
      ProcessValue <- "DIx_DB_M1_QF_Filter_Off_SP"
   Button "Button_9" at 360,10 size 46x20; TextOff 'Inv'
      on Click: InvertBit("DIx_DB_M1_QF_Inverse")
      Appearance <- "DIx_DB_M1_QF_Inverse"
   TextField "Text field_3" at 131,69 size 45x22; Text 'I 0.1'
   TextField "Text field_4" at 176,69 size 120x22; Text 'М2 Готовность'
   Circle "Circle_3" at 131,92 size 22x22
      Appearance <- "DIx_DB_M2_QF_Input"
   Circle "Circle_4" at 154,92 size 22x22
      Appearance <- "DIx_DB_M2_QF_Signal"
   Button "Button_10" at 298,70 size 59x44; TextOff 'Авто'; TextList "Hand"
      on Click: InvertBit("DIx_DB_M2_QF_Hand")
      Appearance <- "DIx_DB_M2_QF_Hand"
      ProcessValue <- "DIx_DB_M2_QF_Hand"
   Button "Button_11" at 240,92 size 49x22; TextOff 'Выкл'
      on Click: ResetBit("DIx_DB_M2_QF_Start_M")
   Button "Button_13" at 184,92 size 47x22; TextOff 'Вкл'
      on Click: SetBit("DIx_DB_M2_QF_Start_M")
      Appearance <- "DIx_DB_M2_QF_Start_M"
   IOField "I/O field_1" at 360,92 size 23x22; FormatPattern 99
      ProcessValue <- "DIx_DB_M2_QF_Filter_On_SP"
   IOField "I/O field_2" at 383,92 size 23x22; FormatPattern 99
      ProcessValue <- "DIx_DB_M2_QF_Filter_Off_SP"
   Button "Button_14" at 360,69 size 46x20; TextOff 'Inv'
      on Click: InvertBit("DIx_DB_M2_QF_Inverse")
      Appearance <- "DIx_DB_M2_QF_Inverse"
   TextField "Text field_5" at 131,128 size 45x22; Text 'I 0.2'
   TextField "Text field_6" at 176,128 size 120x22; Text 'M3 Готовность'
   Circle "Circle_5" at 131,151 size 22x22
      Appearance <- "DIx_DB_M3_QF_Input"
   Circle "Circle_6" at 154,151 size 22x22
      Appearance <- "DIx_DB_M3_QF_Signal"
   Button "Button_15" at 298,129 size 59x44; TextOff 'Авто'; TextList "Hand"
      on Click: InvertBit("DIx_DB_M3_QF_Hand")
      Appearance <- "DIx_DB_M3_QF_Hand"
      ProcessValue <- "DIx_DB_M3_QF_Hand"
   Button "Button_16" at 240,151 size 49x22; TextOff 'Выкл'
      on Click: ResetBit("DIx_DB_M3_QF_Start_M")
   Button "Button_17" at 184,151 size 47x22; TextOff 'Вкл'
      on Click: SetBit("DIx_DB_M3_QF_Start_M")
      Appearance <- "DIx_DB_M3_QF_Start_M"
   IOField "I/O field_3" at 360,151 size 23x22; FormatPattern 99
      ProcessValue <- "DIx_DB_M3_QF_Filter_On_SP"
   IOField "I/O field_4" at 383,151 size 23x22; FormatPattern 99
      ProcessValue <- "DIx_DB_M3_QF_Filter_Off_SP"
   Button "Button_18" at 360,128 size 46x20; TextOff 'Inv'
      on Click: InvertBit("DIx_DB_M3_QF_Inverse")
      Appearance <- "DIx_DB_M3_QF_Inverse"
   TextField "Text field_7" at 131,187 size 45x22; Text 'I 0.3'
   TextField "Text field_8" at 176,187 size 119x22; Text 'Нагреватель 1'
   Circle "Circle_7" at 131,210 size 22x22
      Appearance <- "DIx_DB_Heat_1_Input"
   Circle "Circle_8" at 154,210 size 22x22
      Appearance <- "DIx_DB_Heat_1_Signal"
   Button "Button_19" at 298,188 size 59x44; TextOff 'Авто'; TextList "Hand"
      on Click: InvertBit("DIx_DB_Heat_1_Hand")
      Appearance <- "DIx_DB_Heat_1_Hand"
      ProcessValue <- "DIx_DB_Heat_1_Hand"
   Button "Button_20" at 240,210 size 49x22; TextOff 'Выкл'
      on Click: ResetBit("DIx_DB_Heat_1_Start_M")
   Button "Button_21" at 184,210 size 47x22; TextOff 'Вкл'
      on Click: SetBit("DIx_DB_Heat_1_Start_M")
      Appearance <- "DIx_DB_Heat_1_Start_M"
   IOField "I/O field_5" at 360,210 size 23x22; FormatPattern 99
      ProcessValue <- "DIx_DB_Heat_1_Filter_On_SP"
   IOField "I/O field_8" at 383,210 size 23x22; FormatPattern 99
      ProcessValue <- "DIx_DB_Heat_1_Filter_Off_SP"
   Button "Button_22" at 360,187 size 46x20; TextOff 'Inv'
      on Click: InvertBit("DIx_DB_Heat_1_Inverse")
      Appearance <- "DIx_DB_Heat_1_Inverse"
   TextField "Text field_9" at 131,247 size 45x22; Text 'I 0.4'
   TextField "Text field_10" at 176,247 size 119x22; Text 'Нагреватель 2'
   Circle "Circle_9" at 131,270 size 22x22
      Appearance <- "DIx_DB_Heat_2_Input"
   Circle "Circle_10" at 154,270 size 22x22
      Appearance <- "DIx_DB_Heat_2_Signal"
   Button "Button_23" at 298,248 size 59x44; TextOff 'Авто'; TextList "Hand"
      on Click: InvertBit("DIx_DB_Heat_2_Hand")
      Appearance <- "DIx_DB_Heat_2_Hand"
      ProcessValue <- "DIx_DB_Heat_2_Hand"
   Button "Button_24" at 240,270 size 49x22; TextOff 'Выкл'
      on Click: ResetBit("DIx_DB_Heat_2_Start_M")
   Button "Button_25" at 184,270 size 47x22; TextOff 'Вкл'
      on Click: SetBit("DIx_DB_Heat_2_Start_M")
      Appearance <- "DIx_DB_Heat_2_Start_M"
   IOField "I/O field_9" at 360,270 size 23x22; FormatPattern 99
      ProcessValue <- "DIx_DB_Heat_2_Filter_On_SP"
   IOField "I/O field_10" at 383,270 size 23x22; FormatPattern 99
      ProcessValue <- "DIx_DB_Heat_2_Filter_Off_SP"
   Button "Button_26" at 360,247 size 46x20; TextOff 'Inv'
      on Click: InvertBit("DIx_DB_Heat_2_Inverse")
      Appearance <- "DIx_DB_Heat_2_Inverse"
   TextField "Text field_11" at 131,306 size 45x22; Text 'I 0.5'
   TextField "Text field_12" at 176,306 size 119x22; Text 'Нагреватель 3'
   Circle "Circle_11" at 131,329 size 22x22
      Appearance <- "DIx_DB_Heat_3_Input"
   Circle "Circle_12" at 154,329 size 22x22
      Appearance <- "DIx_DB_Heat_3_Signal"
   Button "Button_27" at 298,307 size 59x44; TextOff 'Авто'; TextList "Hand"
      on Click: InvertBit("DIx_DB_Heat_3_Hand")
      Appearance <- "DIx_DB_Heat_3_Hand"
      ProcessValue <- "DIx_DB_Heat_3_Hand"
   Button "Button_28" at 240,329 size 49x22; TextOff 'Выкл'
      on Click: ResetBit("DIx_DB_Heat_3_Start_M")
   Button "Button_29" at 184,329 size 47x22; TextOff 'Вкл'
      on Click: SetBit("DIx_DB_Heat_3_Start_M")
      Appearance <- "DIx_DB_Heat_3_Start_M"
   IOField "I/O field_11" at 360,329 size 23x22; FormatPattern 99
      ProcessValue <- "DIx_DB_Heat_3_Filter_On_SP"
   IOField "I/O field_12" at 383,329 size 23x22; FormatPattern 99
      ProcessValue <- "DIx_DB_Heat_3_Filter_Off_SP"
   Button "Button_30" at 360,306 size 46x20; TextOff 'Inv'
      on Click: InvertBit("DIx_DB_Heat_3_Inverse")
      Appearance <- "DIx_DB_Heat_3_Inverse"
   TextField "Text field_13" at 131,365 size 45x22; Text 'I 0.6'
   TextField "Text field_14" at 176,365 size 119x22; Text 'Нагреватель 4'
   Circle "Circle_13" at 131,388 size 22x22
      Appearance <- "DIx_DB_Heat_4_Input"
   Circle "Circle_14" at 154,388 size 22x22
      Appearance <- "DIx_DB_Heat_4_Signal"
   Button "Button_31" at 298,366 size 59x44; TextOff 'Авто'; TextList "Hand"
      on Click: InvertBit("DIx_DB_Heat_4_Hand")
      Appearance <- "DIx_DB_Heat_4_Hand"
      ProcessValue <- "DIx_DB_Heat_4_Hand"
   Button "Button_32" at 240,388 size 49x22; TextOff 'Выкл'
      on Click: ResetBit("DIx_DB_Heat_4_Start_M")
   Button "Button_33" at 184,388 size 47x22; TextOff 'Вкл'
      on Click: SetBit("DIx_DB_Heat_4_Start_M")
      Appearance <- "DIx_DB_Heat_4_Start_M"
   IOField "I/O field_13" at 360,388 size 23x22; FormatPattern 99
      ProcessValue <- "DIx_DB_Heat_4_Filter_On_SP"
   IOField "I/O field_14" at 383,388 size 23x22; FormatPattern 99
      ProcessValue <- "DIx_DB_Heat_4_Filter_Off_SP"
   Button "Button_34" at 360,365 size 46x20; TextOff 'Inv'
      on Click: InvertBit("DIx_DB_Heat_4_Inverse")
      Appearance <- "DIx_DB_Heat_4_Inverse"
   TextField "Text field_15" at 131,425 size 45x22; Text 'I 0.7'
   TextField "Text field_16" at 176,425 size 112x22; Text 'Внешний стоп'
   Circle "Circle_15" at 131,448 size 22x22
      Appearance <- "DIx_DB_AllBlock_Input"
   Circle "Circle_16" at 154,448 size 22x22
      Appearance <- "DIx_DB_AllBlock_Signal"
   Button "Button_35" at 298,426 size 59x44; TextOff 'Авто'; TextList "Hand"
      on Click: InvertBit("DIx_DB_AllBlock_Hand")
      Appearance <- "DIx_DB_AllBlock_Hand"
      ProcessValue <- "DIx_DB_AllBlock_Hand"
   Button "Button_36" at 240,448 size 49x22; TextOff 'Выкл'
      on Click: ResetBit("DIx_DB_AllBlock_Start_M")
   Button "Button_37" at 184,448 size 47x22; TextOff 'Вкл'
      on Click: SetBit("DIx_DB_AllBlock_Start_M")
      Appearance <- "DIx_DB_AllBlock_Start_M"
   IOField "I/O field_15" at 360,448 size 23x22; FormatPattern 99
      ProcessValue <- "DIx_DB_AllBlock_Filter_On_SP"
   IOField "I/O field_16" at 383,448 size 23x22; FormatPattern 99
      ProcessValue <- "DIx_DB_AllBlock_Filter_Off_SP"
   Button "Button_38" at 360,425 size 46x20; TextOff 'Inv'
      on Click: InvertBit("DIx_DB_AllBlock_Inverse")
      Appearance <- "DIx_DB_AllBlock_Inverse"
   TextField "Text field_17" at 437,10 size 45x22; Text 'I 1.0'
   TextField "Text field_18" at 482,10 size 59x22; Text 'Весы 1'
   Circle "Circle_17" at 437,33 size 22x22
      Appearance <- "DIx_DB_Mass_1_Input"
   Circle "Circle_18" at 460,33 size 22x22
      Appearance <- "DIx_DB_Mass_1_Signal"
   Button "Button_39" at 604,11 size 59x44; TextOff 'Авто'; TextList "Hand"
      on Click: InvertBit("DIx_DB_Mass_1_Hand")
      Appearance <- "DIx_DB_Mass_1_Hand"
      ProcessValue <- "DIx_DB_Mass_1_Hand"
   Button "Button_40" at 546,33 size 49x22; TextOff 'Выкл'
      on Click: ResetBit("DIx_DB_Mass_1_Start_M")
   Button "Button_41" at 490,33 size 47x22; TextOff 'Вкл'
      on Click: SetBit("DIx_DB_Mass_1_Start_M")
      Appearance <- "DIx_DB_Mass_1_Start_M"
   IOField "I/O field_17" at 666,33 size 23x22; FormatPattern 99
      ProcessValue <- "DIx_DB_Mass_1_Filter_On_SP"
   IOField "I/O field_18" at 689,33 size 23x22; FormatPattern 99
      ProcessValue <- "DIx_DB_Mass_1_Filter_Off_SP"
   Button "Button_42" at 666,10 size 46x20; TextOff 'Inv'
      on Click: InvertBit("DIx_DB_Mass_1_Inverse")
      Appearance <- "DIx_DB_Mass_1_Inverse"
   TextField "Text field_19" at 437,69 size 45x22; Text 'I 1.1'
   TextField "Text field_20" at 482,69 size 59x22; Text 'Весы 2'
   Circle "Circle_19" at 437,92 size 22x22
      Appearance <- "DIx_DB_Mass_2_Input"
   Circle "Circle_20" at 460,92 size 22x22
      Appearance <- "DIx_DB_Mass_2_Signal"
   Button "Button_43" at 604,70 size 59x44; TextOff 'Авто'; TextList "Hand"
      on Click: InvertBit("DIx_DB_Mass_2_Hand")
      Appearance <- "DIx_DB_Mass_2_Hand"
      ProcessValue <- "DIx_DB_Mass_2_Hand"
   Button "Button_44" at 546,92 size 49x22; TextOff 'Выкл'
      on Click: ResetBit("DIx_DB_Mass_2_Start_M")
   Button "Button_45" at 490,92 size 47x22; TextOff 'Вкл'
      on Click: SetBit("DIx_DB_Mass_2_Start_M")
      Appearance <- "DIx_DB_Mass_2_Start_M"
   IOField "I/O field_19" at 666,92 size 23x22; FormatPattern 99
      ProcessValue <- "DIx_DB_Mass_2_Filter_On_SP"
   IOField "I/O field_20" at 689,92 size 23x22; FormatPattern 99
      ProcessValue <- "DIx_DB_Mass_2_Filter_Off_SP"
   Button "Button_46" at 666,69 size 46x20; TextOff 'Inv'
      on Click: InvertBit("DIx_DB_Mass_2_Inverse")